(* Logix 5000 project; controller MV vendor 1 type 14 code 217 rev 31.11; software revision 31.00; part 37 of 53 *)
(* tags used below, declared in another part *)
   MV_Copy_from_fv_file : INT;
   MV_Copy_to_fv_file : INT;
   MV_MV10R : PlantItem;   // MV10R
   MV_MV11R : PlantItem;   // MV11R
   MV_MV12R : PlantItem;   // MV12R
   MV_MV13R : PlantItem;   // MV13R
   MV_MV14R : PlantItem;   // MV14R
   MV_MV15R : PlantItem;   // MV15R
   MV_MV16R : PlantItem;   // MV16R
   MV_MV17R : PlantItem;   // MV17R
   MV_MV18R : PlantItem;   // MV18R
   MV_MV19R : PlantItem;   // MV19R
   MV_MV1R : PlantItem;   // MV1R
   MV_MV20R : PlantItem;   // MV20R
   MV_MV21R : PlantItem;   // MV21R
   MV_MV22R : PlantItem;   // MV22R
   MV_MV23R : PlantItem;   // MV23R
   MV_MV2R : PlantItem;   // MV2R
   MV_MV30R : PlantItem;   // MV30R
   MV_MV31R : PlantItem;   // MV31R
   MV_MV32R : PlantItem;   // MV32R
   MV_MV33R : PlantItem;   // MV33R
   MV_MV34R : PlantItem;   // MV34R
   MV_MV35R : PlantItem;   // MV35R
   MV_MV3R : PlantItem;   // MV3R
   MV_MV4R : PlantItem;   // MV4R
   MV_MV5R : PlantItem;   // MV5R
   MV_MV6R : PlantItem;   // MV6R
   MV_MV7R : PlantItem;   // MV7R
   MV_MV8R : PlantItem;   // MV8R
   MV_MV9R : PlantItem;   // MV9R
   MV_N106 : INT[255];   // ROUSE_BUFF Rouser control vesse l data buffer
   MV_N110 : INT[255];   // MV DATA 0 CURRENT FV DATA
   MV_N111 : INT[50];   // MV 1, CURRENT FV DATA
   MV_N112 : INT[50];   // MV 2, CURRENT FV DATA
   MV_N113 : INT[50];   // MV 3, CURRENT FV DATA
   MV_N114 : INT[50];   // MV 4, CURRENT FV DATA
   MV_N115 : INT[50];   // MV 5, CURRENT FV DATA
   MV_N116 : INT[50];   // MV 6, CURRENT FV DATA
   MV_N117 : INT[50];   // MV 7, CURRENT FV DATA
   MV_N118 : INT[50];   // MV 8, CURRENT FV DATA
   MV_N119 : INT[50];   // MV 9, CURRENT FV DATA
   MV_N120 : INT[50];   // MV 10, CURRENT FV DATA
   MV_N121 : INT[50];   // MV 11, CURRENT FV DATA
   MV_N122 : INT[50];   // MV 12, CURRENT FV DATA
   MV_N123 : INT[50];   // MV 13, CURRENT FV DATA
   MV_N124 : INT[50];   // MV 14, CURRENT FV DATA
   MV_N125 : INT[50];   // MV 15, CURRENT FV DATA
   MV_N126 : INT[50];   // MV 16, CURRENT FV DATA
   MV_N127 : INT[50];   // MV 17, CURRENT FV DATA
   MV_N128 : INT[50];   // MV 18, CURRENT FV DATA
   MV_N129 : INT[50];   // MV 19, CURRENT FV DATA
   MV_N130 : INT[50];   // MV 30, CURRENT FV DATA
   MV_N131 : INT[50];   // MV 31, CURRENT FV DATA
   MV_N132 : INT[50];   // MV 32, CURRENT FV DATA
   MV_N133 : INT[50];   // MV 33, CURRENT FV DATA
   MV_N134 : INT[50];   // MV 34, CURRENT FV DATA
   MV_N135 : INT[50];   // MV 35, CURRENT FV DATA
   MV_N136 : INT[50];   // MV 20, CURRENT FV DATA
   MV_N137 : INT[50];   // MV 21, CURRENT FV DATA
   MV_N138 : INT[50];   // MV 22, CURRENT FV DATA
   MV_N139 : INT[50];   // MV 23, CURRENT FV DATA
   MV_N140 : INT[50];   // MV 36, CURRENT FV DATA
   MV_N141 : INT[50];   // MV 37, CURRENT FV DATA
   MV_N142 : INT[50];   // MV 38, CURRENT FV DATA
   MV_N143 : INT[50];   // MV 39, CURRENT FV DATA
   MV_N144 : INT[50];   // MV 40, CURRENT FV DATA
   MV_N145 : INT[50];   // MV 41, CURRENT FV DATA
   MV_N146 : INT[50];   // MV 42, CURRENT FV DATA
   MV_N147 : INT[50];   // MV 43, CURRENT FV DATA
   MV_N148 : INT[50];   // MV 44, CURRENT FV DATA
   MV_N149 : INT[50];   // MV 45, CURRENT FV DATA
   MV_N150 : INT[50];   // MV 36, CURRENT FV DATA
   MV_N151 : INT[50];   // MV 47, CURRENT FV DATA
   MV_N190 : INT[255];   // Original N File From SLC, No Description Available
(* MV_Common, continued *)

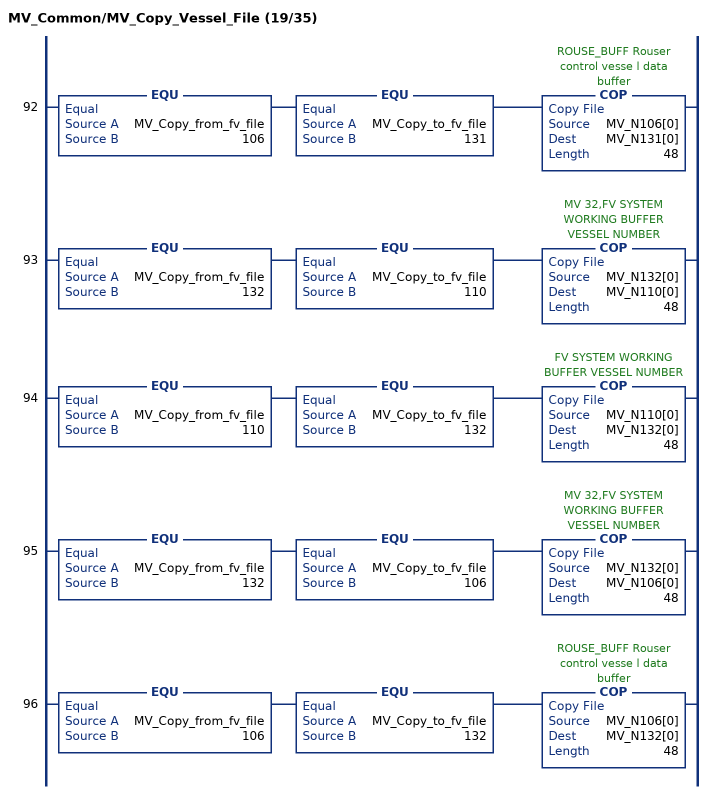
   [picture p861: MV_Common/MV_Copy_Vessel_File rungs 92-96]
   92: EQU(MV_Copy_from_fv_file,106)EQU(MV_Copy_to_fv_file,131)COP(MV_N106[0],MV_N131[0],48);
   93: EQU(MV_Copy_from_fv_file,132)EQU(MV_Copy_to_fv_file,110)COP(MV_N132[0],MV_N110[0],48);
   94: EQU(MV_Copy_from_fv_file,110)EQU(MV_Copy_to_fv_file,132)COP(MV_N110[0],MV_N132[0],48);
   95: EQU(MV_Copy_from_fv_file,132)EQU(MV_Copy_to_fv_file,106)COP(MV_N132[0],MV_N106[0],48);
   96: EQU(MV_Copy_from_fv_file,106)EQU(MV_Copy_to_fv_file,132)COP(MV_N106[0],MV_N132[0],48);
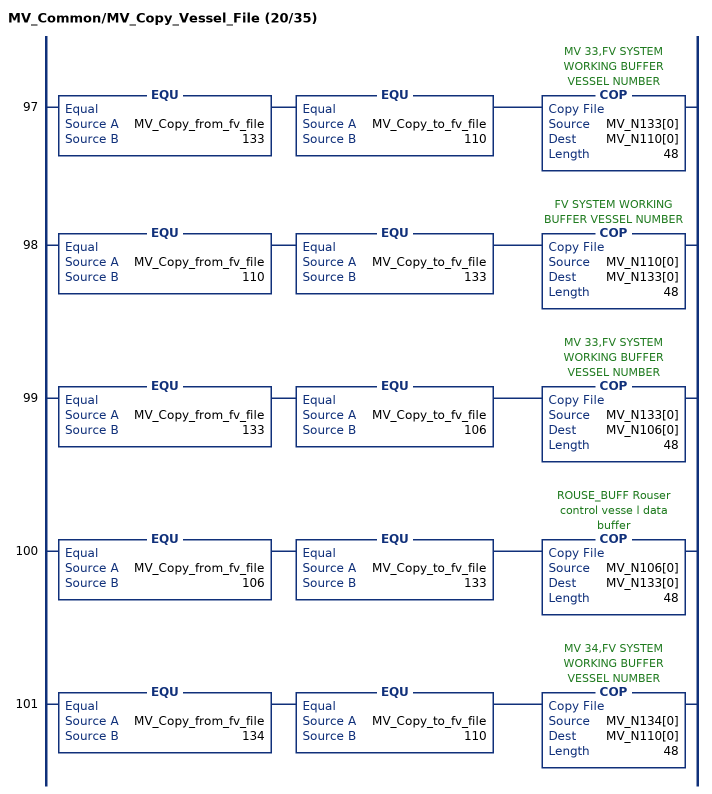
   97: EQU(MV_Copy_from_fv_file,133)EQU(MV_Copy_to_fv_file,110)COP(MV_N133[0],MV_N110[0],48);
   98: EQU(MV_Copy_from_fv_file,110)EQU(MV_Copy_to_fv_file,133)COP(MV_N110[0],MV_N133[0],48);
   99: EQU(MV_Copy_from_fv_file,133)EQU(MV_Copy_to_fv_file,106)COP(MV_N133[0],MV_N106[0],48);
   100: EQU(MV_Copy_from_fv_file,106)EQU(MV_Copy_to_fv_file,133)COP(MV_N106[0],MV_N133[0],48);
   101: EQU(MV_Copy_from_fv_file,134)EQU(MV_Copy_to_fv_file,110)COP(MV_N134[0],MV_N110[0],48);
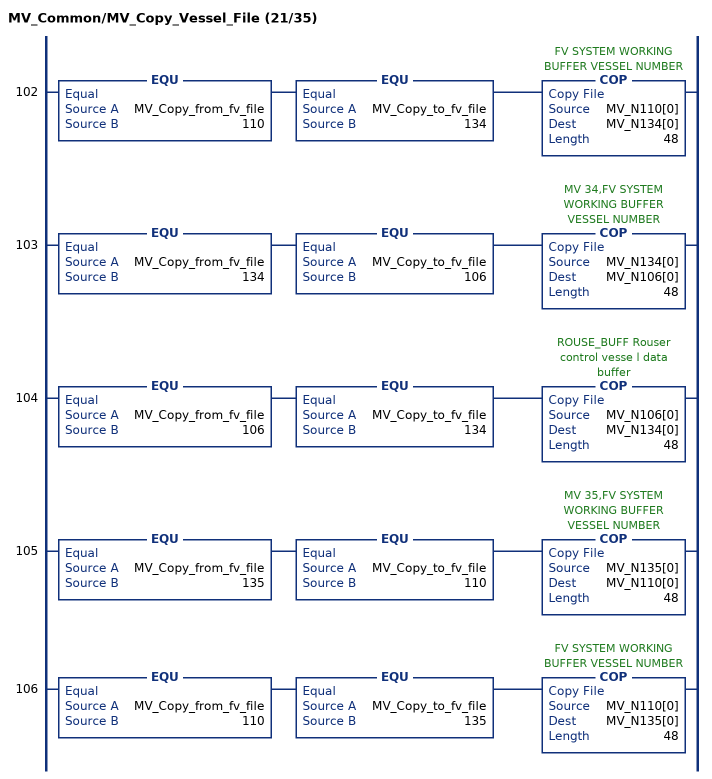
   102: EQU(MV_Copy_from_fv_file,110)EQU(MV_Copy_to_fv_file,134)COP(MV_N110[0],MV_N134[0],48);
   103: EQU(MV_Copy_from_fv_file,134)EQU(MV_Copy_to_fv_file,106)COP(MV_N134[0],MV_N106[0],48);
   104: EQU(MV_Copy_from_fv_file,106)EQU(MV_Copy_to_fv_file,134)COP(MV_N106[0],MV_N134[0],48);
   105: EQU(MV_Copy_from_fv_file,135)EQU(MV_Copy_to_fv_file,110)COP(MV_N135[0],MV_N110[0],48);
   106: EQU(MV_Copy_from_fv_file,110)EQU(MV_Copy_to_fv_file,135)COP(MV_N110[0],MV_N135[0],48);
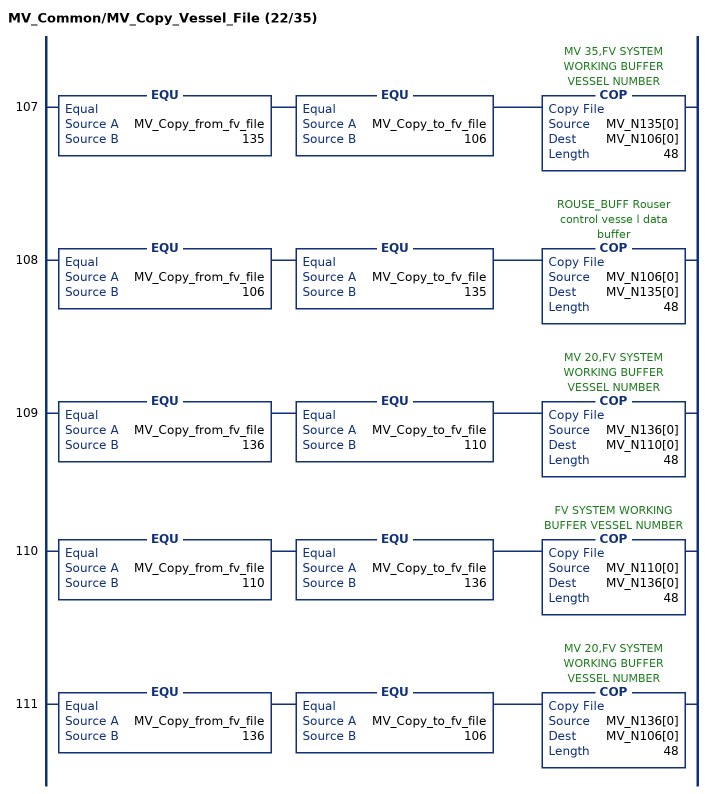
   107: EQU(MV_Copy_from_fv_file,135)EQU(MV_Copy_to_fv_file,106)COP(MV_N135[0],MV_N106[0],48);
   108: EQU(MV_Copy_from_fv_file,106)EQU(MV_Copy_to_fv_file,135)COP(MV_N106[0],MV_N135[0],48);
   109: EQU(MV_Copy_from_fv_file,136)EQU(MV_Copy_to_fv_file,110)COP(MV_N136[0],MV_N110[0],48);
   110: EQU(MV_Copy_from_fv_file,110)EQU(MV_Copy_to_fv_file,136)COP(MV_N110[0],MV_N136[0],48);
   111: EQU(MV_Copy_from_fv_file,136)EQU(MV_Copy_to_fv_file,106)COP(MV_N136[0],MV_N106[0],48);
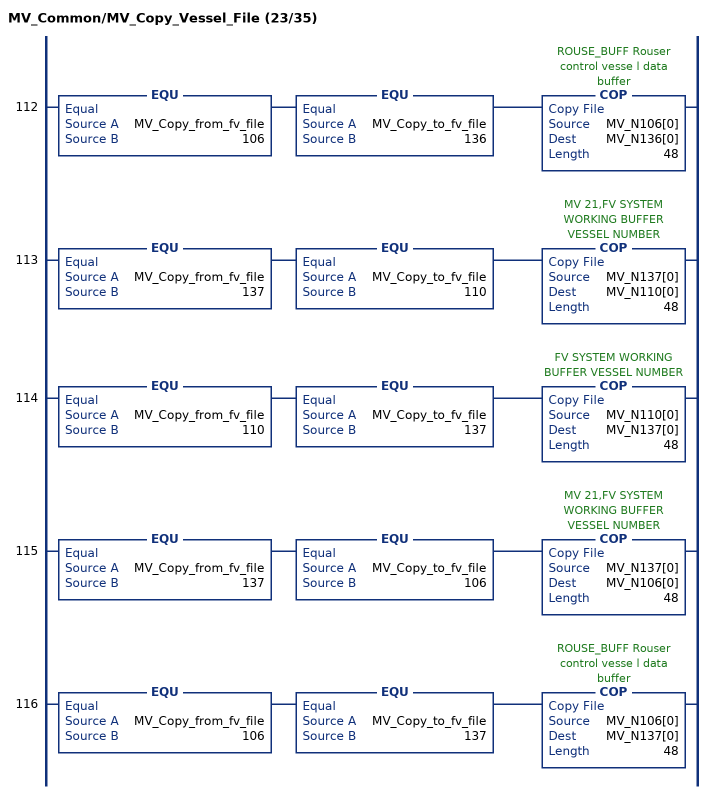
   112: EQU(MV_Copy_from_fv_file,106)EQU(MV_Copy_to_fv_file,136)COP(MV_N106[0],MV_N136[0],48);
   113: EQU(MV_Copy_from_fv_file,137)EQU(MV_Copy_to_fv_file,110)COP(MV_N137[0],MV_N110[0],48);
   114: EQU(MV_Copy_from_fv_file,110)EQU(MV_Copy_to_fv_file,137)COP(MV_N110[0],MV_N137[0],48);
   115: EQU(MV_Copy_from_fv_file,137)EQU(MV_Copy_to_fv_file,106)COP(MV_N137[0],MV_N106[0],48);
   116: EQU(MV_Copy_from_fv_file,106)EQU(MV_Copy_to_fv_file,137)COP(MV_N106[0],MV_N137[0],48);
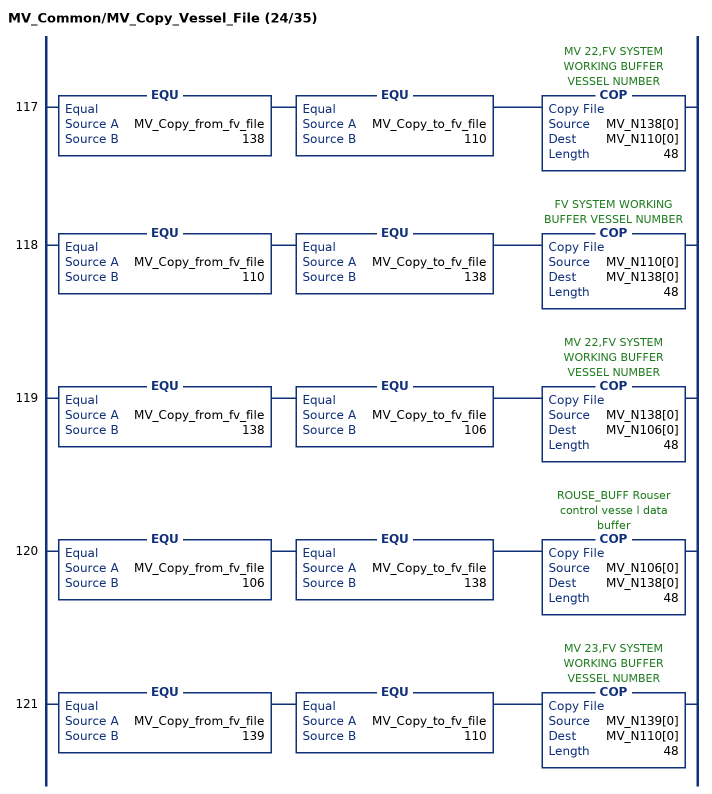
   117: EQU(MV_Copy_from_fv_file,138)EQU(MV_Copy_to_fv_file,110)COP(MV_N138[0],MV_N110[0],48);
   118: EQU(MV_Copy_from_fv_file,110)EQU(MV_Copy_to_fv_file,138)COP(MV_N110[0],MV_N138[0],48);
   119: EQU(MV_Copy_from_fv_file,138)EQU(MV_Copy_to_fv_file,106)COP(MV_N138[0],MV_N106[0],48);
   120: EQU(MV_Copy_from_fv_file,106)EQU(MV_Copy_to_fv_file,138)COP(MV_N106[0],MV_N138[0],48);
   121: EQU(MV_Copy_from_fv_file,139)EQU(MV_Copy_to_fv_file,110)COP(MV_N139[0],MV_N110[0],48);
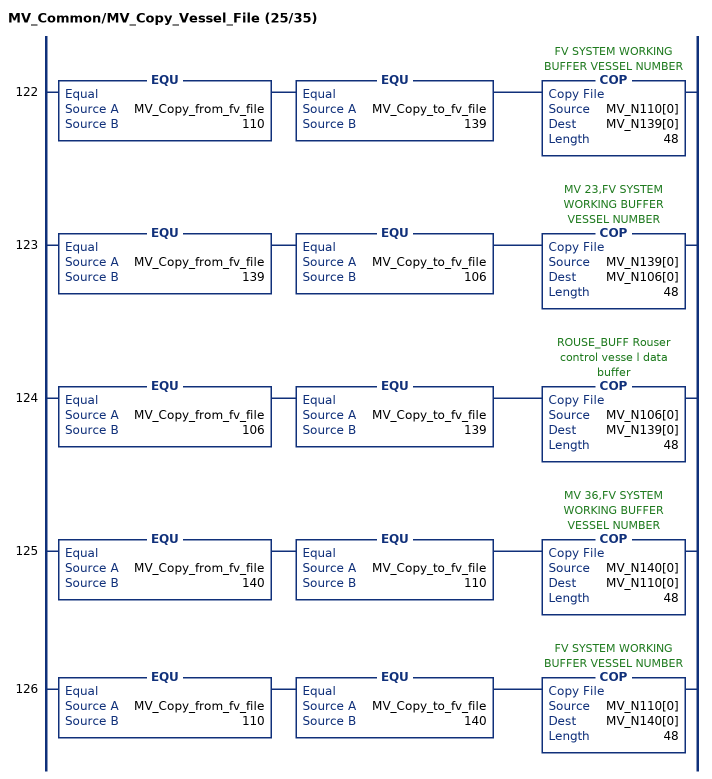
   122: EQU(MV_Copy_from_fv_file,110)EQU(MV_Copy_to_fv_file,139)COP(MV_N110[0],MV_N139[0],48);
   123: EQU(MV_Copy_from_fv_file,139)EQU(MV_Copy_to_fv_file,106)COP(MV_N139[0],MV_N106[0],48);
   124: EQU(MV_Copy_from_fv_file,106)EQU(MV_Copy_to_fv_file,139)COP(MV_N106[0],MV_N139[0],48);
   125: EQU(MV_Copy_from_fv_file,140)EQU(MV_Copy_to_fv_file,110)COP(MV_N140[0],MV_N110[0],48);
   126: EQU(MV_Copy_from_fv_file,110)EQU(MV_Copy_to_fv_file,140)COP(MV_N110[0],MV_N140[0],48);
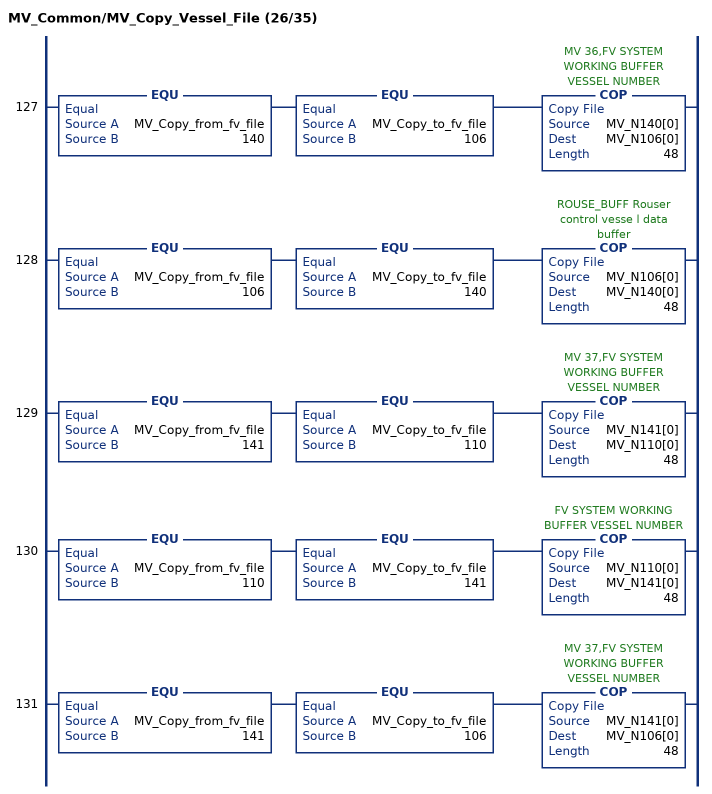
   127: EQU(MV_Copy_from_fv_file,140)EQU(MV_Copy_to_fv_file,106)COP(MV_N140[0],MV_N106[0],48);
   128: EQU(MV_Copy_from_fv_file,106)EQU(MV_Copy_to_fv_file,140)COP(MV_N106[0],MV_N140[0],48);
   129: EQU(MV_Copy_from_fv_file,141)EQU(MV_Copy_to_fv_file,110)COP(MV_N141[0],MV_N110[0],48);
   130: EQU(MV_Copy_from_fv_file,110)EQU(MV_Copy_to_fv_file,141)COP(MV_N110[0],MV_N141[0],48);
   131: EQU(MV_Copy_from_fv_file,141)EQU(MV_Copy_to_fv_file,106)COP(MV_N141[0],MV_N106[0],48);
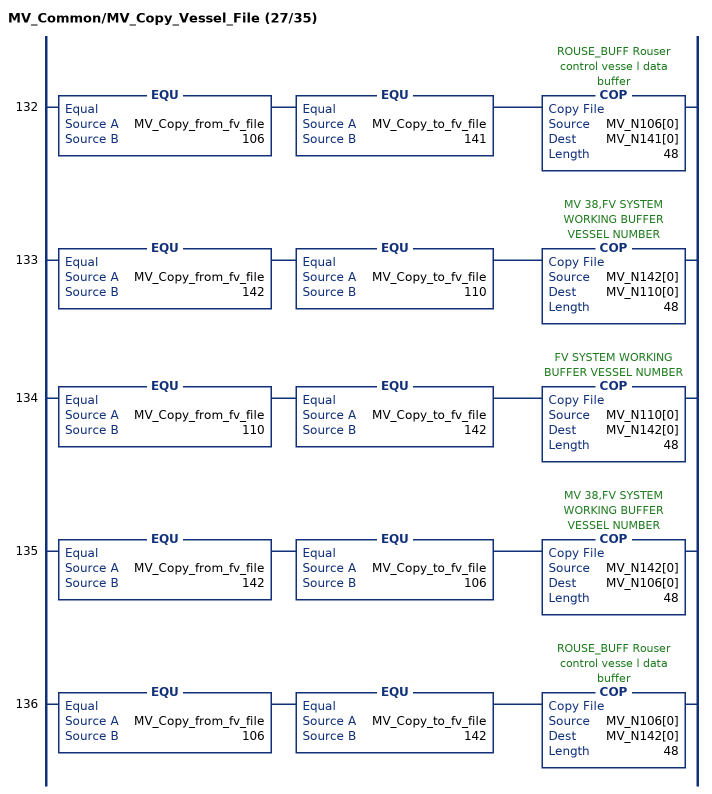
   132: EQU(MV_Copy_from_fv_file,106)EQU(MV_Copy_to_fv_file,141)COP(MV_N106[0],MV_N141[0],48);
   133: EQU(MV_Copy_from_fv_file,142)EQU(MV_Copy_to_fv_file,110)COP(MV_N142[0],MV_N110[0],48);
   134: EQU(MV_Copy_from_fv_file,110)EQU(MV_Copy_to_fv_file,142)COP(MV_N110[0],MV_N142[0],48);
   135: EQU(MV_Copy_from_fv_file,142)EQU(MV_Copy_to_fv_file,106)COP(MV_N142[0],MV_N106[0],48);
   136: EQU(MV_Copy_from_fv_file,106)EQU(MV_Copy_to_fv_file,142)COP(MV_N106[0],MV_N142[0],48);
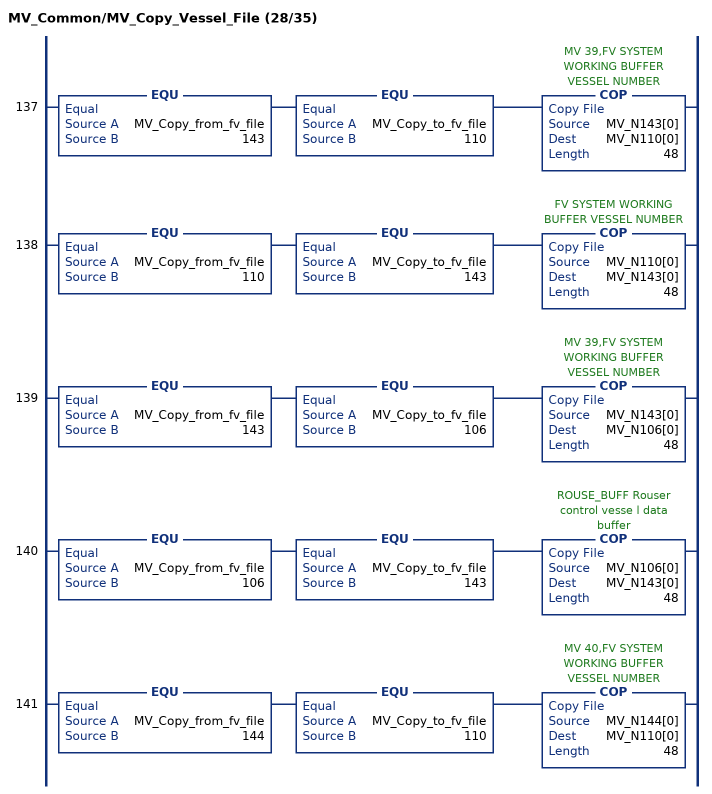
   137: EQU(MV_Copy_from_fv_file,143)EQU(MV_Copy_to_fv_file,110)COP(MV_N143[0],MV_N110[0],48);
   138: EQU(MV_Copy_from_fv_file,110)EQU(MV_Copy_to_fv_file,143)COP(MV_N110[0],MV_N143[0],48);
   139: EQU(MV_Copy_from_fv_file,143)EQU(MV_Copy_to_fv_file,106)COP(MV_N143[0],MV_N106[0],48);
   140: EQU(MV_Copy_from_fv_file,106)EQU(MV_Copy_to_fv_file,143)COP(MV_N106[0],MV_N143[0],48);
   141: EQU(MV_Copy_from_fv_file,144)EQU(MV_Copy_to_fv_file,110)COP(MV_N144[0],MV_N110[0],48);
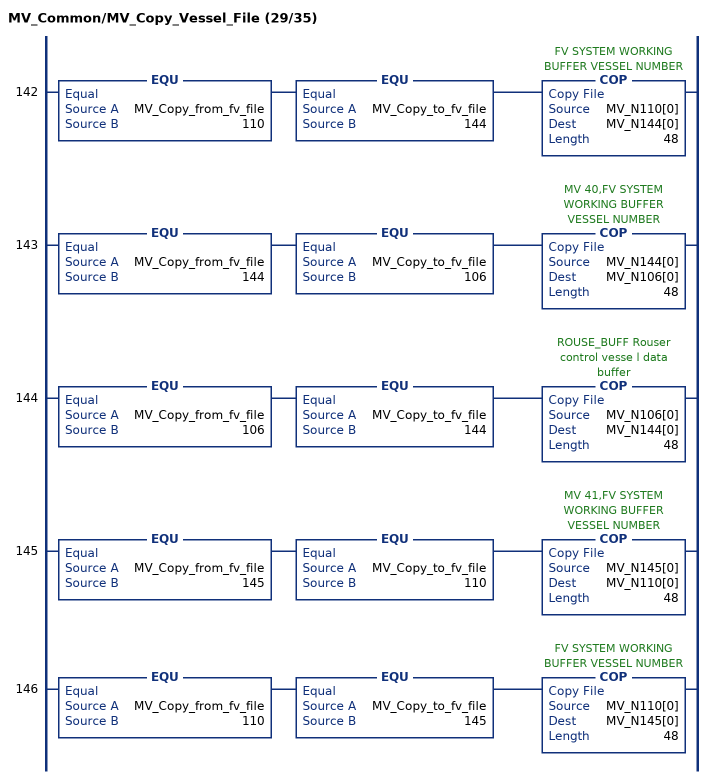
   142: EQU(MV_Copy_from_fv_file,110)EQU(MV_Copy_to_fv_file,144)COP(MV_N110[0],MV_N144[0],48);
   143: EQU(MV_Copy_from_fv_file,144)EQU(MV_Copy_to_fv_file,106)COP(MV_N144[0],MV_N106[0],48);
   144: EQU(MV_Copy_from_fv_file,106)EQU(MV_Copy_to_fv_file,144)COP(MV_N106[0],MV_N144[0],48);
   145: EQU(MV_Copy_from_fv_file,145)EQU(MV_Copy_to_fv_file,110)COP(MV_N145[0],MV_N110[0],48);
   146: EQU(MV_Copy_from_fv_file,110)EQU(MV_Copy_to_fv_file,145)COP(MV_N110[0],MV_N145[0],48);
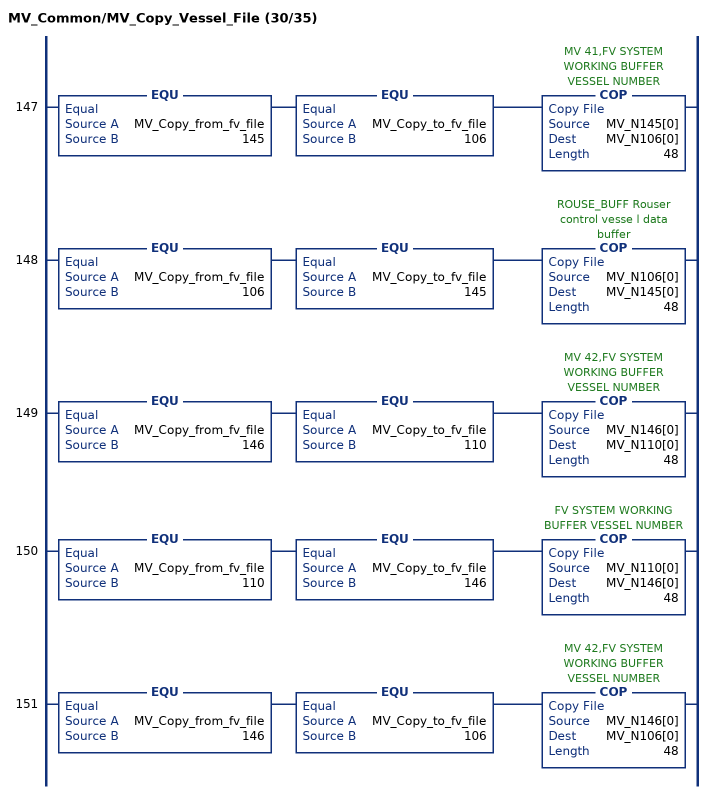
   147: EQU(MV_Copy_from_fv_file,145)EQU(MV_Copy_to_fv_file,106)COP(MV_N145[0],MV_N106[0],48);
   148: EQU(MV_Copy_from_fv_file,106)EQU(MV_Copy_to_fv_file,145)COP(MV_N106[0],MV_N145[0],48);
   149: EQU(MV_Copy_from_fv_file,146)EQU(MV_Copy_to_fv_file,110)COP(MV_N146[0],MV_N110[0],48);
   150: EQU(MV_Copy_from_fv_file,110)EQU(MV_Copy_to_fv_file,146)COP(MV_N110[0],MV_N146[0],48);
   151: EQU(MV_Copy_from_fv_file,146)EQU(MV_Copy_to_fv_file,106)COP(MV_N146[0],MV_N106[0],48);
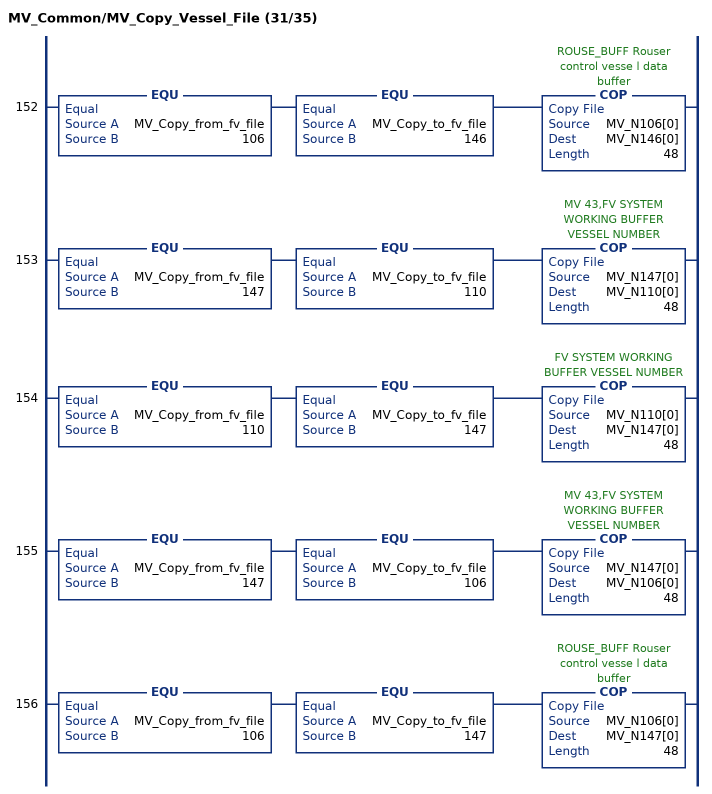
   152: EQU(MV_Copy_from_fv_file,106)EQU(MV_Copy_to_fv_file,146)COP(MV_N106[0],MV_N146[0],48);
   153: EQU(MV_Copy_from_fv_file,147)EQU(MV_Copy_to_fv_file,110)COP(MV_N147[0],MV_N110[0],48);
   154: EQU(MV_Copy_from_fv_file,110)EQU(MV_Copy_to_fv_file,147)COP(MV_N110[0],MV_N147[0],48);
   155: EQU(MV_Copy_from_fv_file,147)EQU(MV_Copy_to_fv_file,106)COP(MV_N147[0],MV_N106[0],48);
   156: EQU(MV_Copy_from_fv_file,106)EQU(MV_Copy_to_fv_file,147)COP(MV_N106[0],MV_N147[0],48);
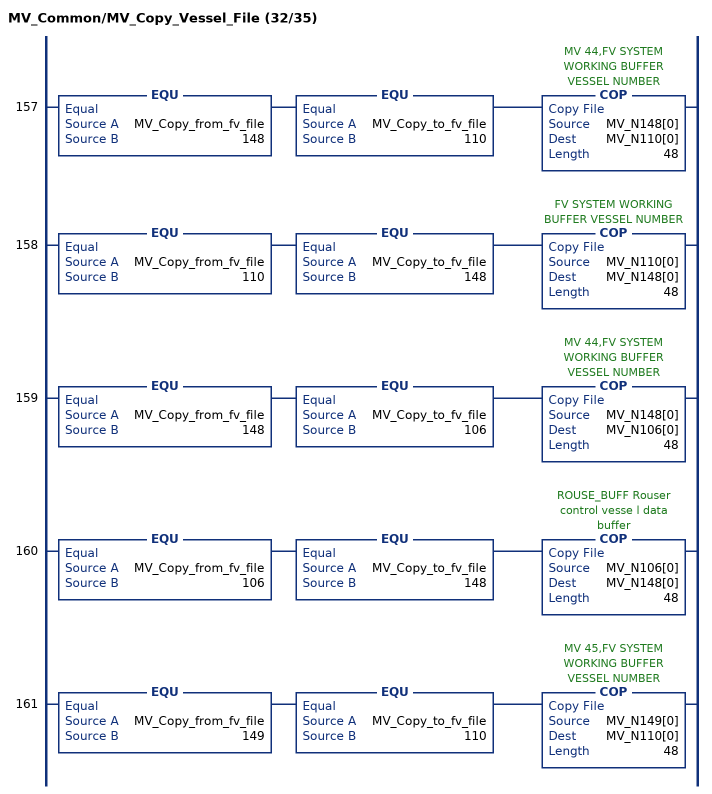
   157: EQU(MV_Copy_from_fv_file,148)EQU(MV_Copy_to_fv_file,110)COP(MV_N148[0],MV_N110[0],48);
   158: EQU(MV_Copy_from_fv_file,110)EQU(MV_Copy_to_fv_file,148)COP(MV_N110[0],MV_N148[0],48);
   159: EQU(MV_Copy_from_fv_file,148)EQU(MV_Copy_to_fv_file,106)COP(MV_N148[0],MV_N106[0],48);
   160: EQU(MV_Copy_from_fv_file,106)EQU(MV_Copy_to_fv_file,148)COP(MV_N106[0],MV_N148[0],48);
   161: EQU(MV_Copy_from_fv_file,149)EQU(MV_Copy_to_fv_file,110)COP(MV_N149[0],MV_N110[0],48);
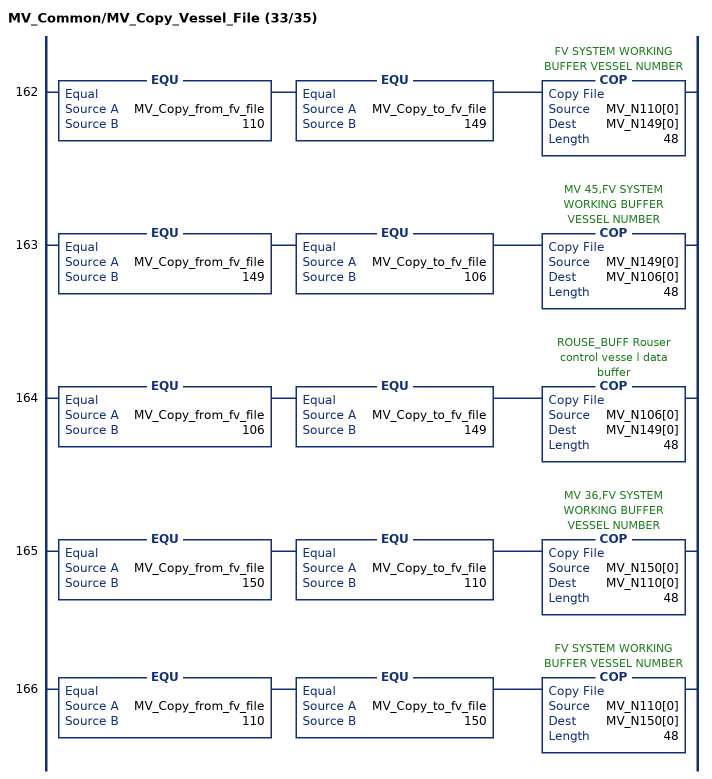
   162: EQU(MV_Copy_from_fv_file,110)EQU(MV_Copy_to_fv_file,149)COP(MV_N110[0],MV_N149[0],48);
   163: EQU(MV_Copy_from_fv_file,149)EQU(MV_Copy_to_fv_file,106)COP(MV_N149[0],MV_N106[0],48);
   164: EQU(MV_Copy_from_fv_file,106)EQU(MV_Copy_to_fv_file,149)COP(MV_N106[0],MV_N149[0],48);
   165: EQU(MV_Copy_from_fv_file,150)EQU(MV_Copy_to_fv_file,110)COP(MV_N150[0],MV_N110[0],48);
   166: EQU(MV_Copy_from_fv_file,110)EQU(MV_Copy_to_fv_file,150)COP(MV_N110[0],MV_N150[0],48);
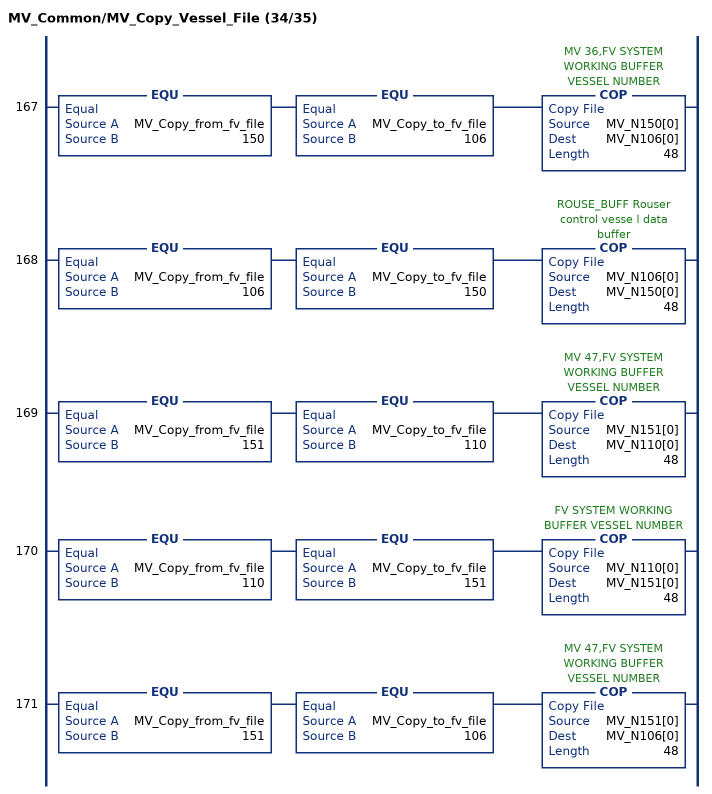
   167: EQU(MV_Copy_from_fv_file,150)EQU(MV_Copy_to_fv_file,106)COP(MV_N150[0],MV_N106[0],48);
   168: EQU(MV_Copy_from_fv_file,106)EQU(MV_Copy_to_fv_file,150)COP(MV_N106[0],MV_N150[0],48);
   169: EQU(MV_Copy_from_fv_file,151)EQU(MV_Copy_to_fv_file,110)COP(MV_N151[0],MV_N110[0],48);
   170: EQU(MV_Copy_from_fv_file,110)EQU(MV_Copy_to_fv_file,151)COP(MV_N110[0],MV_N151[0],48);
   171: EQU(MV_Copy_from_fv_file,151)EQU(MV_Copy_to_fv_file,106)COP(MV_N151[0],MV_N106[0],48);
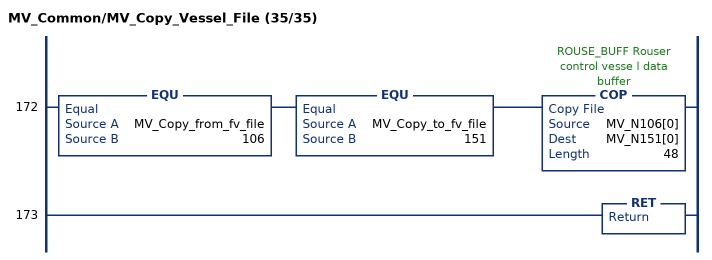
   172: EQU(MV_Copy_from_fv_file,106)EQU(MV_Copy_to_fv_file,151)COP(MV_N106[0],MV_N151[0],48);
   173: RET();
END_ROUTINE

ROUTINE MV_DIG_OUTPUT_6   (* ladder *)
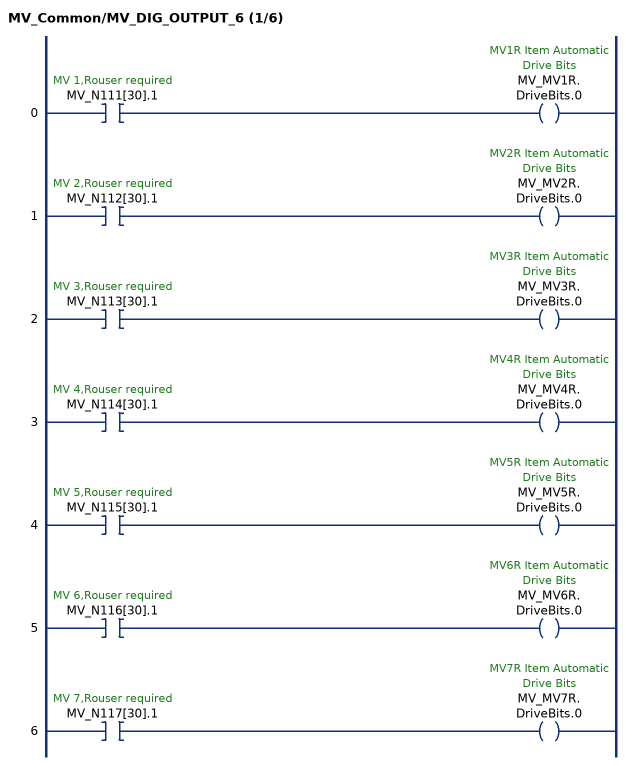
   0: XIC(MV_N111[30].1)OTE(MV_MV1R.DriveBits.0);
   1: XIC(MV_N112[30].1)OTE(MV_MV2R.DriveBits.0);
   2: XIC(MV_N113[30].1)OTE(MV_MV3R.DriveBits.0);
   3: XIC(MV_N114[30].1)OTE(MV_MV4R.DriveBits.0);
   4: XIC(MV_N115[30].1)OTE(MV_MV5R.DriveBits.0);
   5: XIC(MV_N116[30].1)OTE(MV_MV6R.DriveBits.0);
   6: XIC(MV_N117[30].1)OTE(MV_MV7R.DriveBits.0);
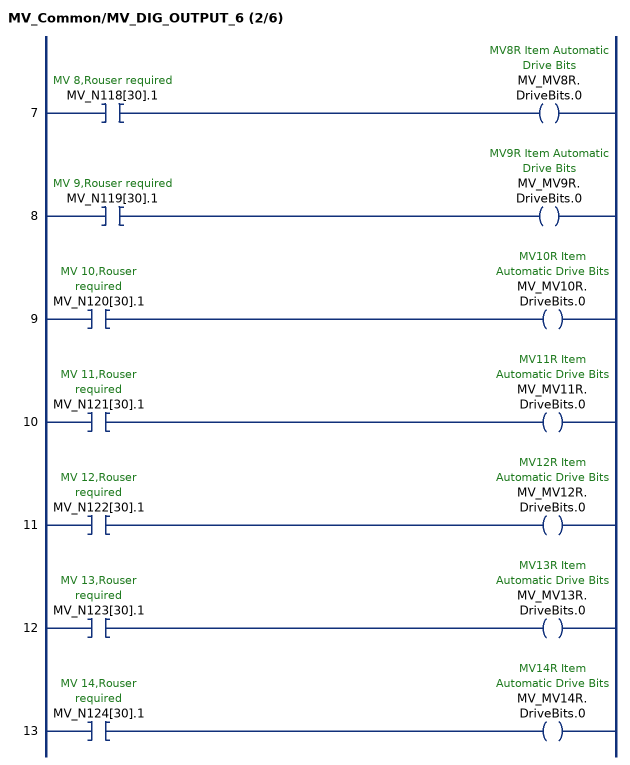
   7: XIC(MV_N118[30].1)OTE(MV_MV8R.DriveBits.0);
   8: XIC(MV_N119[30].1)OTE(MV_MV9R.DriveBits.0);
   9: XIC(MV_N120[30].1)OTE(MV_MV10R.DriveBits.0);
   10: XIC(MV_N121[30].1)OTE(MV_MV11R.DriveBits.0);
   11: XIC(MV_N122[30].1)OTE(MV_MV12R.DriveBits.0);
   12: XIC(MV_N123[30].1)OTE(MV_MV13R.DriveBits.0);
   13: XIC(MV_N124[30].1)OTE(MV_MV14R.DriveBits.0);
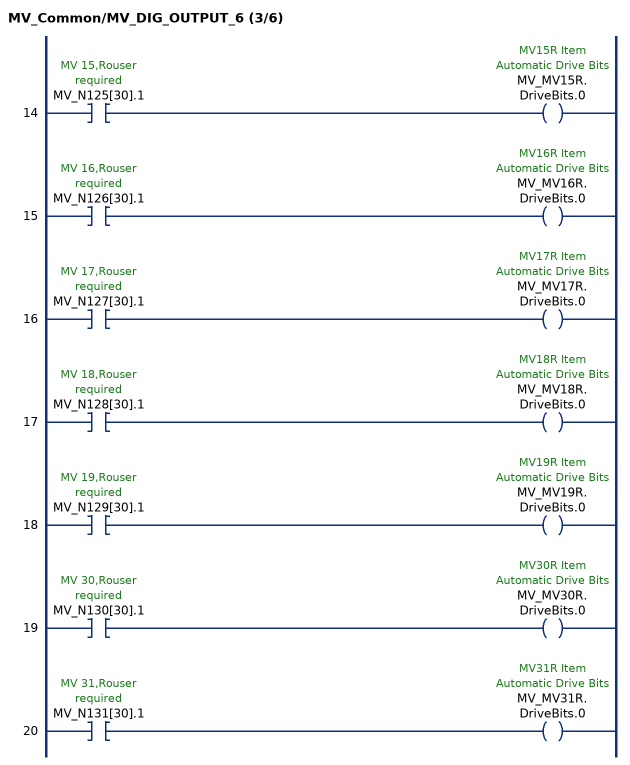
   14: XIC(MV_N125[30].1)OTE(MV_MV15R.DriveBits.0);
   15: XIC(MV_N126[30].1)OTE(MV_MV16R.DriveBits.0);
   16: XIC(MV_N127[30].1)OTE(MV_MV17R.DriveBits.0);
   17: XIC(MV_N128[30].1)OTE(MV_MV18R.DriveBits.0);
   18: XIC(MV_N129[30].1)OTE(MV_MV19R.DriveBits.0);
   19: XIC(MV_N130[30].1)OTE(MV_MV30R.DriveBits.0);
   20: XIC(MV_N131[30].1)OTE(MV_MV31R.DriveBits.0);
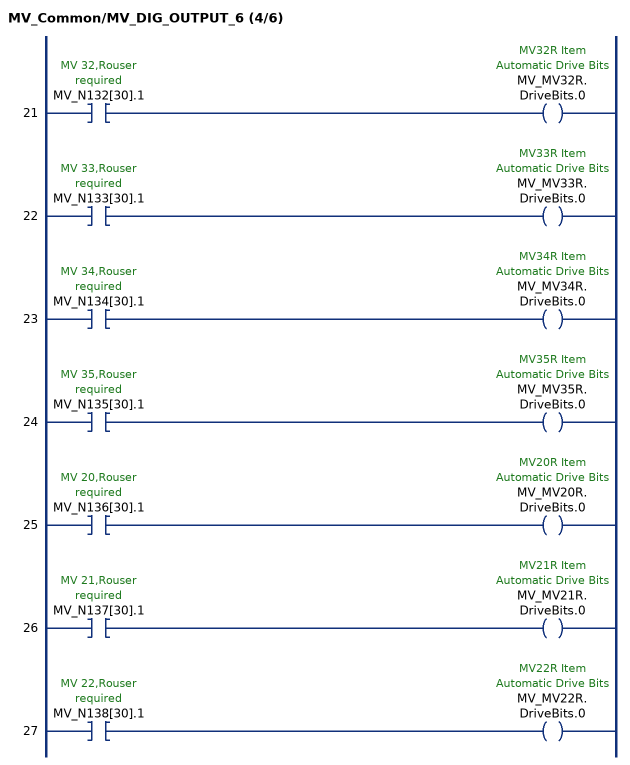
   21: XIC(MV_N132[30].1)OTE(MV_MV32R.DriveBits.0);
   22: XIC(MV_N133[30].1)OTE(MV_MV33R.DriveBits.0);
   23: XIC(MV_N134[30].1)OTE(MV_MV34R.DriveBits.0);
   24: XIC(MV_N135[30].1)OTE(MV_MV35R.DriveBits.0);
   25: XIC(MV_N136[30].1)OTE(MV_MV20R.DriveBits.0);
   26: XIC(MV_N137[30].1)OTE(MV_MV21R.DriveBits.0);
   27: XIC(MV_N138[30].1)OTE(MV_MV22R.DriveBits.0);
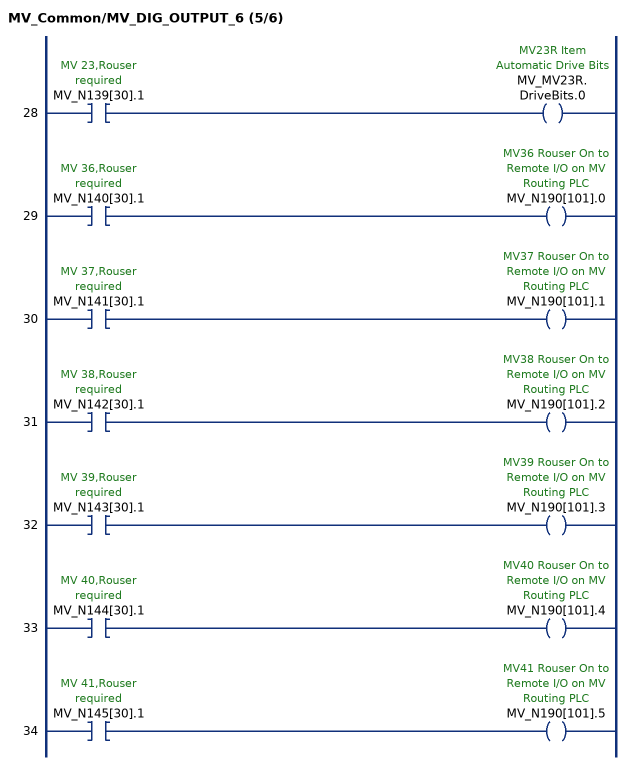
   28: XIC(MV_N139[30].1)OTE(MV_MV23R.DriveBits.0);
   29: XIC(MV_N140[30].1)OTE(MV_N190[101].0);
   30: XIC(MV_N141[30].1)OTE(MV_N190[101].1);
   31: XIC(MV_N142[30].1)OTE(MV_N190[101].2);
   32: XIC(MV_N143[30].1)OTE(MV_N190[101].3);
   33: XIC(MV_N144[30].1)OTE(MV_N190[101].4);
   34: XIC(MV_N145[30].1)OTE(MV_N190[101].5);
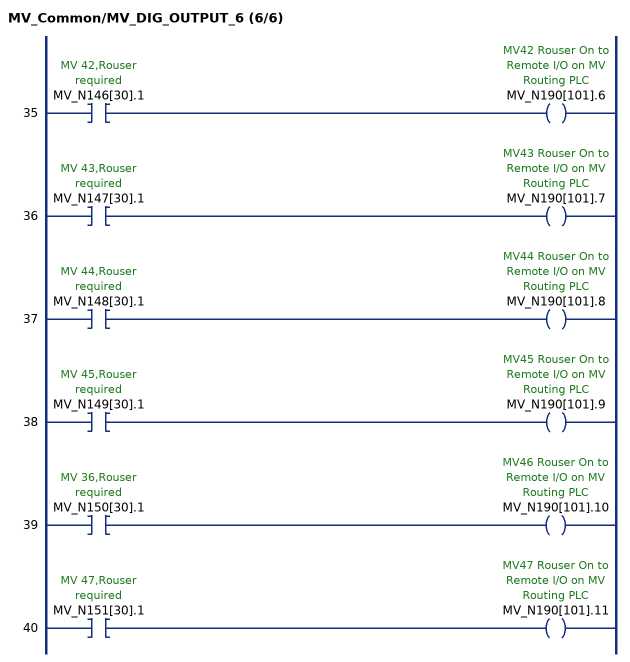
   35: XIC(MV_N146[30].1)OTE(MV_N190[101].6);
   36: XIC(MV_N147[30].1)OTE(MV_N190[101].7);
   37: XIC(MV_N148[30].1)OTE(MV_N190[101].8);
   38: XIC(MV_N149[30].1)OTE(MV_N190[101].9);
   39: XIC(MV_N150[30].1)OTE(MV_N190[101].10);
   40: XIC(MV_N151[30].1)OTE(MV_N190[101].11);
END_ROUTINE
